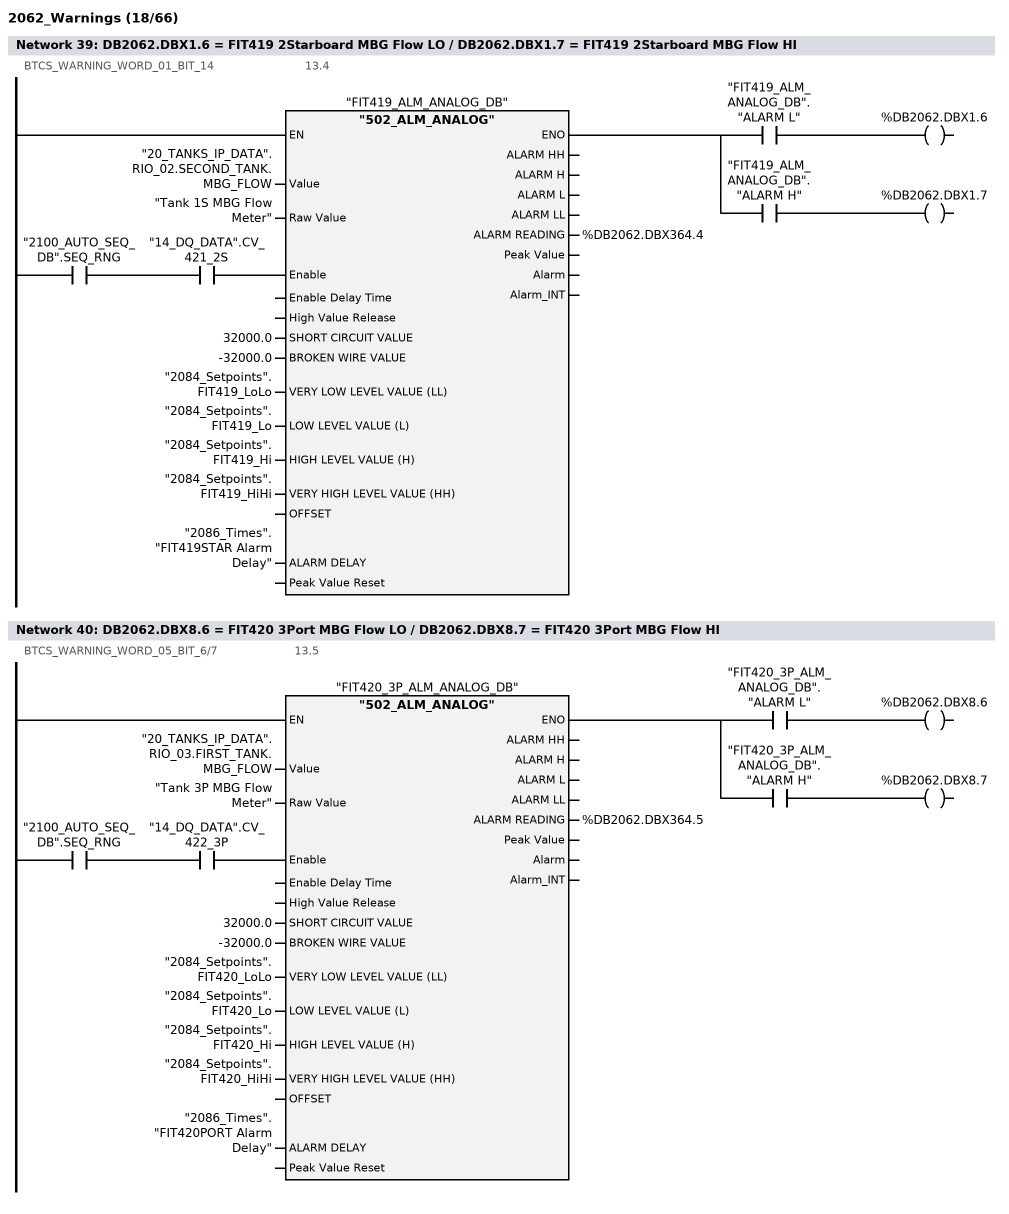
   RUNG wire#powerrail
      "FIT419_ALM_ANALOG_DB"(Enable := wire#w1, Value := "20_TANKS_IP_DATA".RIO_02.SECOND_TANK.MBG_FLOW, "Raw Value" := "Tank 1S MBG Flow Meter", "Enable Delay Time" :=, "High Value Release" :=, "SHORT CIRCUIT VALUE" := 32000.0, "BROKEN WIRE VALUE" := -32000.0, "VERY LOW LEVEL VALUE (LL)" := "2084_Setpoints".FIT419_LoLo, "LOW LEVEL VALUE (L)" := "2084_Setpoints".FIT419_Lo, "HIGH LEVEL VALUE (H)" := "2084_Setpoints".FIT419_Hi, "VERY HIGH LEVEL VALUE (HH)" := "2084_Setpoints".FIT419_HiHi, OFFSET :=, "ALARM DELAY" := "2086_Times"."FIT419STAR Alarm Delay", "Peak Value Reset" :=, "ALARM HH" =>, "ALARM H" =>, "ALARM L" =>, "ALARM LL" =>, "ALARM READING" => %DB2062.DBX364.4, "Peak Value" =>, Alarm =>, Alarm_INT =>)
      wire#w2
      Contact( "FIT419_ALM_ANALOG_DB"."ALARM L" )
      Coil( %DB2062.DBX1.6 )
   END_RUNG
   RUNG wire#powerrail
      Contact( "2100_AUTO_SEQ_DB".SEQ_RNG )
      Contact( "14_DQ_DATA".CV_421_2S )
   END_RUNG wire#w1
   RUNG wire#w2
      Contact( "FIT419_ALM_ANALOG_DB"."ALARM H" )
      Coil( %DB2062.DBX1.7 )
   END_RUNG
   // the same network as SCL:
   "FIT419_ALM_ANALOG_DB"(Value := "20_TANKS_IP_DATA".RIO_02.SECOND_TANK.MBG_FLOW,   // "502_ALM_ANALOG"
                          "Raw Value" := "Tank 1S MBG Flow Meter",
                          Enable := "2100_AUTO_SEQ_DB".SEQ_RNG AND "14_DQ_DATA".CV_421_2S,
                          "SHORT CIRCUIT VALUE" := 32000.0,
                          "BROKEN WIRE VALUE" := -32000.0,
                          "VERY LOW LEVEL VALUE (LL)" := "2084_Setpoints".FIT419_LoLo,
                          "LOW LEVEL VALUE (L)" := "2084_Setpoints".FIT419_Lo,
                          "HIGH LEVEL VALUE (H)" := "2084_Setpoints".FIT419_Hi,
                          "VERY HIGH LEVEL VALUE (HH)" := "2084_Setpoints".FIT419_HiHi,
                          "ALARM DELAY" := "2086_Times"."FIT419STAR Alarm Delay",
                          "ALARM READING" => %DB2062.DBX364.4,
                          ENO => #_w1);
   %DB2062.DBX1.6 := #_w1 AND "FIT419_ALM_ANALOG_DB"."ALARM L";
   %DB2062.DBX1.7 := #_w1 AND "FIT419_ALM_ANALOG_DB"."ALARM H";
END_REGION

REGION Network 40: DB2062.DBX8.6 = FIT420 3Port MBG Flow LO / DB2062.DBX8.7 = FIT420 3Port MBG Flow HI
   // BTCS_WARNING_WORD_05_BIT_6/7                      13.5
   RUNG wire#powerrail
      "FIT420_3P_ALM_ANALOG_DB"(Enable := wire#w1, Value := "20_TANKS_IP_DATA".RIO_03.FIRST_TANK.MBG_FLOW, "Raw Value" := "Tank 3P MBG Flow Meter", "Enable Delay Time" :=, "High Value Release" :=, "SHORT CIRCUIT VALUE" := 32000.0, "BROKEN WIRE VALUE" := -32000.0, "VERY LOW LEVEL VALUE (LL)" := "2084_Setpoints".FIT420_LoLo, "LOW LEVEL VALUE (L)" := "2084_Setpoints".FIT420_Lo, "HIGH LEVEL VALUE (H)" := "2084_Setpoints".FIT420_Hi, "VERY HIGH LEVEL VALUE (HH)" := "2084_Setpoints".FIT420_HiHi, OFFSET :=, "ALARM DELAY" := "2086_Times"."FIT420PORT Alarm Delay", "Peak Value Reset" :=, "ALARM HH" =>, "ALARM H" =>, "ALARM L" =>, "ALARM LL" =>, "ALARM READING" => %DB2062.DBX364.5, "Peak Value" =>, Alarm =>, Alarm_INT =>)
      wire#w2
      Contact( "FIT420_3P_ALM_ANALOG_DB"."ALARM L" )
      Coil( %DB2062.DBX8.6 )
   END_RUNG
   RUNG wire#powerrail
      Contact( "2100_AUTO_SEQ_DB".SEQ_RNG )
      Contact( "14_DQ_DATA".CV_422_3P )
   END_RUNG wire#w1
   RUNG wire#w2
      Contact( "FIT420_3P_ALM_ANALOG_DB"."ALARM H" )
      Coil( %DB2062.DBX8.7 )
   END_RUNG
   // the same network as SCL:
   "FIT420_3P_ALM_ANALOG_DB"(Value := "20_TANKS_IP_DATA".RIO_03.FIRST_TANK.MBG_FLOW,   // "502_ALM_ANALOG"
                           "Raw Value" := "Tank 3P MBG Flow Meter",
                           Enable := "2100_AUTO_SEQ_DB".SEQ_RNG AND "14_DQ_DATA".CV_422_3P,
                           "SHORT CIRCUIT VALUE" := 32000.0,
                           "BROKEN WIRE VALUE" := -32000.0,
                           "VERY LOW LEVEL VALUE (LL)" := "2084_Setpoints".FIT420_LoLo,
                           "LOW LEVEL VALUE (L)" := "2084_Setpoints".FIT420_Lo,
                           "HIGH LEVEL VALUE (H)" := "2084_Setpoints".FIT420_Hi,
                           "VERY HIGH LEVEL VALUE (HH)" := "2084_Setpoints".FIT420_HiHi,
                           "ALARM DELAY" := "2086_Times"."FIT420PORT Alarm Delay",
                           "ALARM READING" => %DB2062.DBX364.5,
                           ENO => #_w1);
   %DB2062.DBX8.6 := #_w1 AND "FIT420_3P_ALM_ANALOG_DB"."ALARM L";
   %DB2062.DBX8.7 := #_w1 AND "FIT420_3P_ALM_ANALOG_DB"."ALARM H";
END_REGION

REGION Network 41: DB2062.DBX9.0 = FIT419 3Starboard MBG Flow LO / DB2062.DBX9.1 = FIT419 3Starboard MBG Flow HI
   // BTCS_WARNING_WORD_05_BIT_8/9                13.6
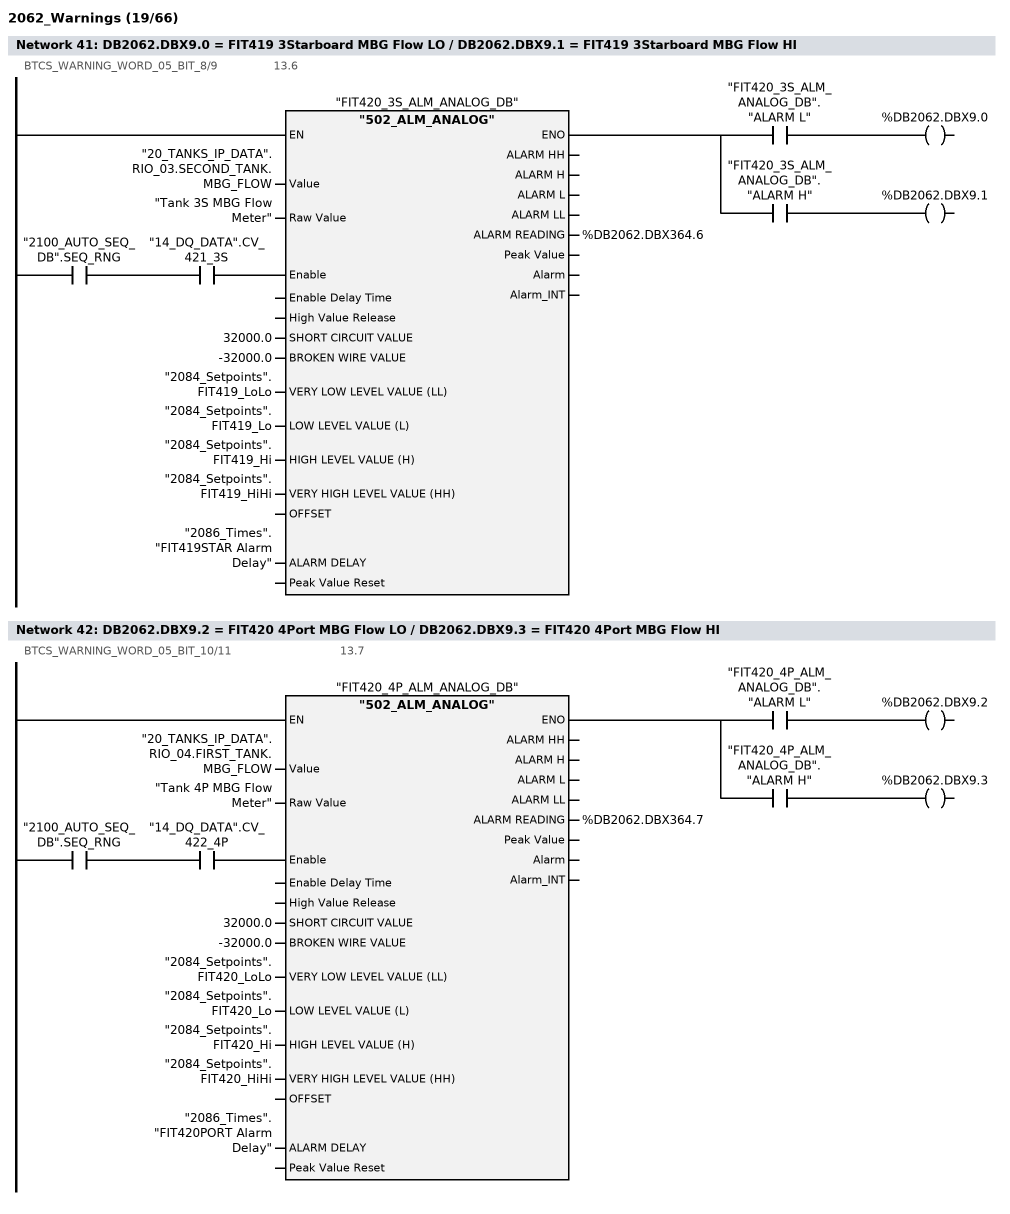
   RUNG wire#powerrail
      "FIT420_3S_ALM_ANALOG_DB"(Enable := wire#w1, Value := "20_TANKS_IP_DATA".RIO_03.SECOND_TANK.MBG_FLOW, "Raw Value" := "Tank 3S MBG Flow Meter", "Enable Delay Time" :=, "High Value Release" :=, "SHORT CIRCUIT VALUE" := 32000.0, "BROKEN WIRE VALUE" := -32000.0, "VERY LOW LEVEL VALUE (LL)" := "2084_Setpoints".FIT419_LoLo, "LOW LEVEL VALUE (L)" := "2084_Setpoints".FIT419_Lo, "HIGH LEVEL VALUE (H)" := "2084_Setpoints".FIT419_Hi, "VERY HIGH LEVEL VALUE (HH)" := "2084_Setpoints".FIT419_HiHi, OFFSET :=, "ALARM DELAY" := "2086_Times"."FIT419STAR Alarm Delay", "Peak Value Reset" :=, "ALARM HH" =>, "ALARM H" =>, "ALARM L" =>, "ALARM LL" =>, "ALARM READING" => %DB2062.DBX364.6, "Peak Value" =>, Alarm =>, Alarm_INT =>)
      wire#w2
      Contact( "FIT420_3S_ALM_ANALOG_DB"."ALARM L" )
      Coil( %DB2062.DBX9.0 )
   END_RUNG
   RUNG wire#powerrail
      Contact( "2100_AUTO_SEQ_DB".SEQ_RNG )
      Contact( "14_DQ_DATA".CV_421_3S )
   END_RUNG wire#w1
   RUNG wire#w2
      Contact( "FIT420_3S_ALM_ANALOG_DB"."ALARM H" )
      Coil( %DB2062.DBX9.1 )
   END_RUNG
   // the same network as SCL:
   "FIT420_3S_ALM_ANALOG_DB"(Value := "20_TANKS_IP_DATA".RIO_03.SECOND_TANK.MBG_FLOW,   // "502_ALM_ANALOG"
                           "Raw Value" := "Tank 3S MBG Flow Meter",
                           Enable := "2100_AUTO_SEQ_DB".SEQ_RNG AND "14_DQ_DATA".CV_421_3S,
                           "SHORT CIRCUIT VALUE" := 32000.0,
                           "BROKEN WIRE VALUE" := -32000.0,
                           "VERY LOW LEVEL VALUE (LL)" := "2084_Setpoints".FIT419_LoLo,
                           "LOW LEVEL VALUE (L)" := "2084_Setpoints".FIT419_Lo,
                           "HIGH LEVEL VALUE (H)" := "2084_Setpoints".FIT419_Hi,
                           "VERY HIGH LEVEL VALUE (HH)" := "2084_Setpoints".FIT419_HiHi,
                           "ALARM DELAY" := "2086_Times"."FIT419STAR Alarm Delay",
                           "ALARM READING" => %DB2062.DBX364.6,
                           ENO => #_w1);
   %DB2062.DBX9.0 := #_w1 AND "FIT420_3S_ALM_ANALOG_DB"."ALARM L";
   %DB2062.DBX9.1 := #_w1 AND "FIT420_3S_ALM_ANALOG_DB"."ALARM H";
END_REGION

REGION Network 42: DB2062.DBX9.2 = FIT420 4Port MBG Flow LO / DB2062.DBX9.3 = FIT420 4Port MBG Flow HI
   // BTCS_WARNING_WORD_05_BIT_10/11                               13.7
   RUNG wire#powerrail
      "FIT420_4P_ALM_ANALOG_DB"(Enable := wire#w1, Value := "20_TANKS_IP_DATA".RIO_04.FIRST_TANK.MBG_FLOW, "Raw Value" := "Tank 4P MBG Flow Meter", "Enable Delay Time" :=, "High Value Release" :=, "SHORT CIRCUIT VALUE" := 32000.0, "BROKEN WIRE VALUE" := -32000.0, "VERY LOW LEVEL VALUE (LL)" := "2084_Setpoints".FIT420_LoLo, "LOW LEVEL VALUE (L)" := "2084_Setpoints".FIT420_Lo, "HIGH LEVEL VALUE (H)" := "2084_Setpoints".FIT420_Hi, "VERY HIGH LEVEL VALUE (HH)" := "2084_Setpoints".FIT420_HiHi, OFFSET :=, "ALARM DELAY" := "2086_Times"."FIT420PORT Alarm Delay", "Peak Value Reset" :=, "ALARM HH" =>, "ALARM H" =>, "ALARM L" =>, "ALARM LL" =>, "ALARM READING" => %DB2062.DBX364.7, "Peak Value" =>, Alarm =>, Alarm_INT =>)
      wire#w2
      Contact( "FIT420_4P_ALM_ANALOG_DB"."ALARM L" )
      Coil( %DB2062.DBX9.2 )
   END_RUNG
   RUNG wire#powerrail
      Contact( "2100_AUTO_SEQ_DB".SEQ_RNG )
      Contact( "14_DQ_DATA".CV_422_4P )
   END_RUNG wire#w1
   RUNG wire#w2
      Contact( "FIT420_4P_ALM_ANALOG_DB"."ALARM H" )
      Coil( %DB2062.DBX9.3 )
   END_RUNG
   // the same network as SCL:
   "FIT420_4P_ALM_ANALOG_DB"(Value := "20_TANKS_IP_DATA".RIO_04.FIRST_TANK.MBG_FLOW,   // "502_ALM_ANALOG"
                           "Raw Value" := "Tank 4P MBG Flow Meter",
                           Enable := "2100_AUTO_SEQ_DB".SEQ_RNG AND "14_DQ_DATA".CV_422_4P,
                           "SHORT CIRCUIT VALUE" := 32000.0,
                           "BROKEN WIRE VALUE" := -32000.0,
                           "VERY LOW LEVEL VALUE (LL)" := "2084_Setpoints".FIT420_LoLo,
                           "LOW LEVEL VALUE (L)" := "2084_Setpoints".FIT420_Lo,
                           "HIGH LEVEL VALUE (H)" := "2084_Setpoints".FIT420_Hi,
                           "VERY HIGH LEVEL VALUE (HH)" := "2084_Setpoints".FIT420_HiHi,
                           "ALARM DELAY" := "2086_Times"."FIT420PORT Alarm Delay",
                           "ALARM READING" => %DB2062.DBX364.7,
                           ENO => #_w1);
   %DB2062.DBX9.2 := #_w1 AND "FIT420_4P_ALM_ANALOG_DB"."ALARM L";
   %DB2062.DBX9.3 := #_w1 AND "FIT420_4P_ALM_ANALOG_DB"."ALARM H";
END_REGION

REGION Network 43: DB2062.DBX9.4 = FIT419 4Starboard MBG Flow LO / DB2062.DBX9.5 = FIT419 4Starboard MBG Flow HI
   // BTCS_WARNING_WORD_05_BIT_12/13                               13.8
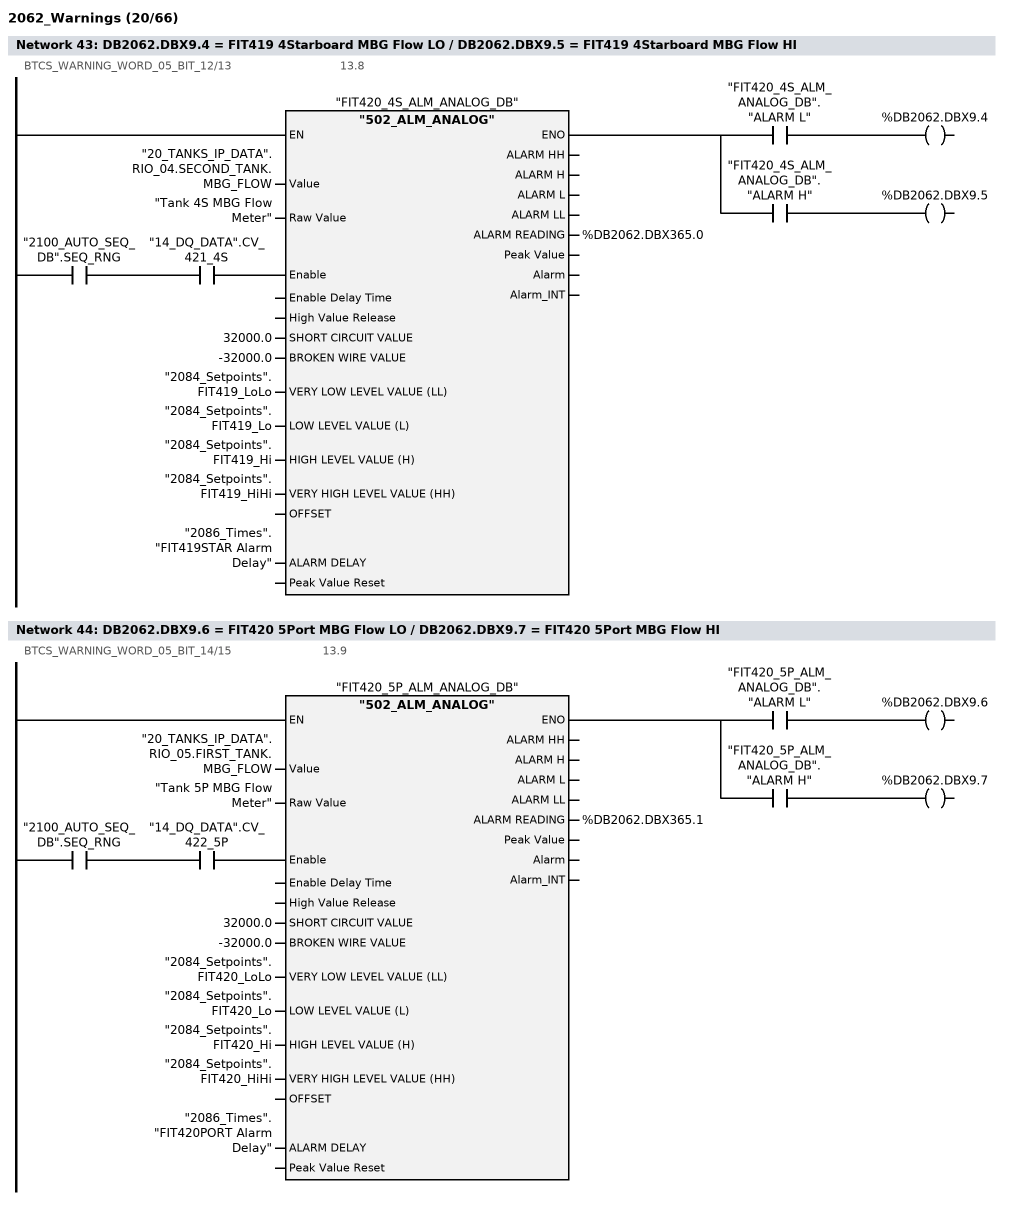
   RUNG wire#powerrail
      "FIT420_4S_ALM_ANALOG_DB"(Enable := wire#w1, Value := "20_TANKS_IP_DATA".RIO_04.SECOND_TANK.MBG_FLOW, "Raw Value" := "Tank 4S MBG Flow Meter", "Enable Delay Time" :=, "High Value Release" :=, "SHORT CIRCUIT VALUE" := 32000.0, "BROKEN WIRE VALUE" := -32000.0, "VERY LOW LEVEL VALUE (LL)" := "2084_Setpoints".FIT419_LoLo, "LOW LEVEL VALUE (L)" := "2084_Setpoints".FIT419_Lo, "HIGH LEVEL VALUE (H)" := "2084_Setpoints".FIT419_Hi, "VERY HIGH LEVEL VALUE (HH)" := "2084_Setpoints".FIT419_HiHi, OFFSET :=, "ALARM DELAY" := "2086_Times"."FIT419STAR Alarm Delay", "Peak Value Reset" :=, "ALARM HH" =>, "ALARM H" =>, "ALARM L" =>, "ALARM LL" =>, "ALARM READING" => %DB2062.DBX365.0, "Peak Value" =>, Alarm =>, Alarm_INT =>)
      wire#w2
      Contact( "FIT420_4S_ALM_ANALOG_DB"."ALARM L" )
      Coil( %DB2062.DBX9.4 )
   END_RUNG
   RUNG wire#powerrail
      Contact( "2100_AUTO_SEQ_DB".SEQ_RNG )
      Contact( "14_DQ_DATA".CV_421_4S )
   END_RUNG wire#w1
   RUNG wire#w2
      Contact( "FIT420_4S_ALM_ANALOG_DB"."ALARM H" )
      Coil( %DB2062.DBX9.5 )
   END_RUNG
   // the same network as SCL:
   "FIT420_4S_ALM_ANALOG_DB"(Value := "20_TANKS_IP_DATA".RIO_04.SECOND_TANK.MBG_FLOW,   // "502_ALM_ANALOG"
                           "Raw Value" := "Tank 4S MBG Flow Meter",
                           Enable := "2100_AUTO_SEQ_DB".SEQ_RNG AND "14_DQ_DATA".CV_421_4S,
                           "SHORT CIRCUIT VALUE" := 32000.0,
                           "BROKEN WIRE VALUE" := -32000.0,
                           "VERY LOW LEVEL VALUE (LL)" := "2084_Setpoints".FIT419_LoLo,
                           "LOW LEVEL VALUE (L)" := "2084_Setpoints".FIT419_Lo,
                           "HIGH LEVEL VALUE (H)" := "2084_Setpoints".FIT419_Hi,
                           "VERY HIGH LEVEL VALUE (HH)" := "2084_Setpoints".FIT419_HiHi,
                           "ALARM DELAY" := "2086_Times"."FIT419STAR Alarm Delay",
                           "ALARM READING" => %DB2062.DBX365.0,
                           ENO => #_w1);
   %DB2062.DBX9.4 := #_w1 AND "FIT420_4S_ALM_ANALOG_DB"."ALARM L";
   %DB2062.DBX9.5 := #_w1 AND "FIT420_4S_ALM_ANALOG_DB"."ALARM H";
END_REGION

REGION Network 44: DB2062.DBX9.6 = FIT420 5Port MBG Flow LO / DB2062.DBX9.7 = FIT420 5Port MBG Flow HI
   // BTCS_WARNING_WORD_05_BIT_14/15                          13.9
   RUNG wire#powerrail
      "FIT420_5P_ALM_ANALOG_DB"(Enable := wire#w1, Value := "20_TANKS_IP_DATA".RIO_05.FIRST_TANK.MBG_FLOW, "Raw Value" := "Tank 5P MBG Flow Meter", "Enable Delay Time" :=, "High Value Release" :=, "SHORT CIRCUIT VALUE" := 32000.0, "BROKEN WIRE VALUE" := -32000.0, "VERY LOW LEVEL VALUE (LL)" := "2084_Setpoints".FIT420_LoLo, "LOW LEVEL VALUE (L)" := "2084_Setpoints".FIT420_Lo, "HIGH LEVEL VALUE (H)" := "2084_Setpoints".FIT420_Hi, "VERY HIGH LEVEL VALUE (HH)" := "2084_Setpoints".FIT420_HiHi, OFFSET :=, "ALARM DELAY" := "2086_Times"."FIT420PORT Alarm Delay", "Peak Value Reset" :=, "ALARM HH" =>, "ALARM H" =>, "ALARM L" =>, "ALARM LL" =>, "ALARM READING" => %DB2062.DBX365.1, "Peak Value" =>, Alarm =>, Alarm_INT =>)
      wire#w2
      Contact( "FIT420_5P_ALM_ANALOG_DB"."ALARM L" )
      Coil( %DB2062.DBX9.6 )
   END_RUNG
   RUNG wire#powerrail
      Contact( "2100_AUTO_SEQ_DB".SEQ_RNG )
      Contact( "14_DQ_DATA".CV_422_5P )
   END_RUNG wire#w1
   RUNG wire#w2
      Contact( "FIT420_5P_ALM_ANALOG_DB"."ALARM H" )
      Coil( %DB2062.DBX9.7 )
   END_RUNG
   // the same network as SCL:
   "FIT420_5P_ALM_ANALOG_DB"(Value := "20_TANKS_IP_DATA".RIO_05.FIRST_TANK.MBG_FLOW,   // "502_ALM_ANALOG"
                           "Raw Value" := "Tank 5P MBG Flow Meter",
                           Enable := "2100_AUTO_SEQ_DB".SEQ_RNG AND "14_DQ_DATA".CV_422_5P,
                           "SHORT CIRCUIT VALUE" := 32000.0,
                           "BROKEN WIRE VALUE" := -32000.0,
                           "VERY LOW LEVEL VALUE (LL)" := "2084_Setpoints".FIT420_LoLo,
                           "LOW LEVEL VALUE (L)" := "2084_Setpoints".FIT420_Lo,
                           "HIGH LEVEL VALUE (H)" := "2084_Setpoints".FIT420_Hi,
                           "VERY HIGH LEVEL VALUE (HH)" := "2084_Setpoints".FIT420_HiHi,
                           "ALARM DELAY" := "2086_Times"."FIT420PORT Alarm Delay",
                           "ALARM READING" => %DB2062.DBX365.1,
                           ENO => #_w1);
   %DB2062.DBX9.6 := #_w1 AND "FIT420_5P_ALM_ANALOG_DB"."ALARM L";
   %DB2062.DBX9.7 := #_w1 AND "FIT420_5P_ALM_ANALOG_DB"."ALARM H";
END_REGION

REGION Network 45: DB2062.DBX10.0 = FIT419 5Starboard MBG Flow LO / DB2062.DBX10.1 = FIT419 5Starboard MBG Flow HI
   // BTCS_WARNING_WORD_06_BIT_0/1                         13.10
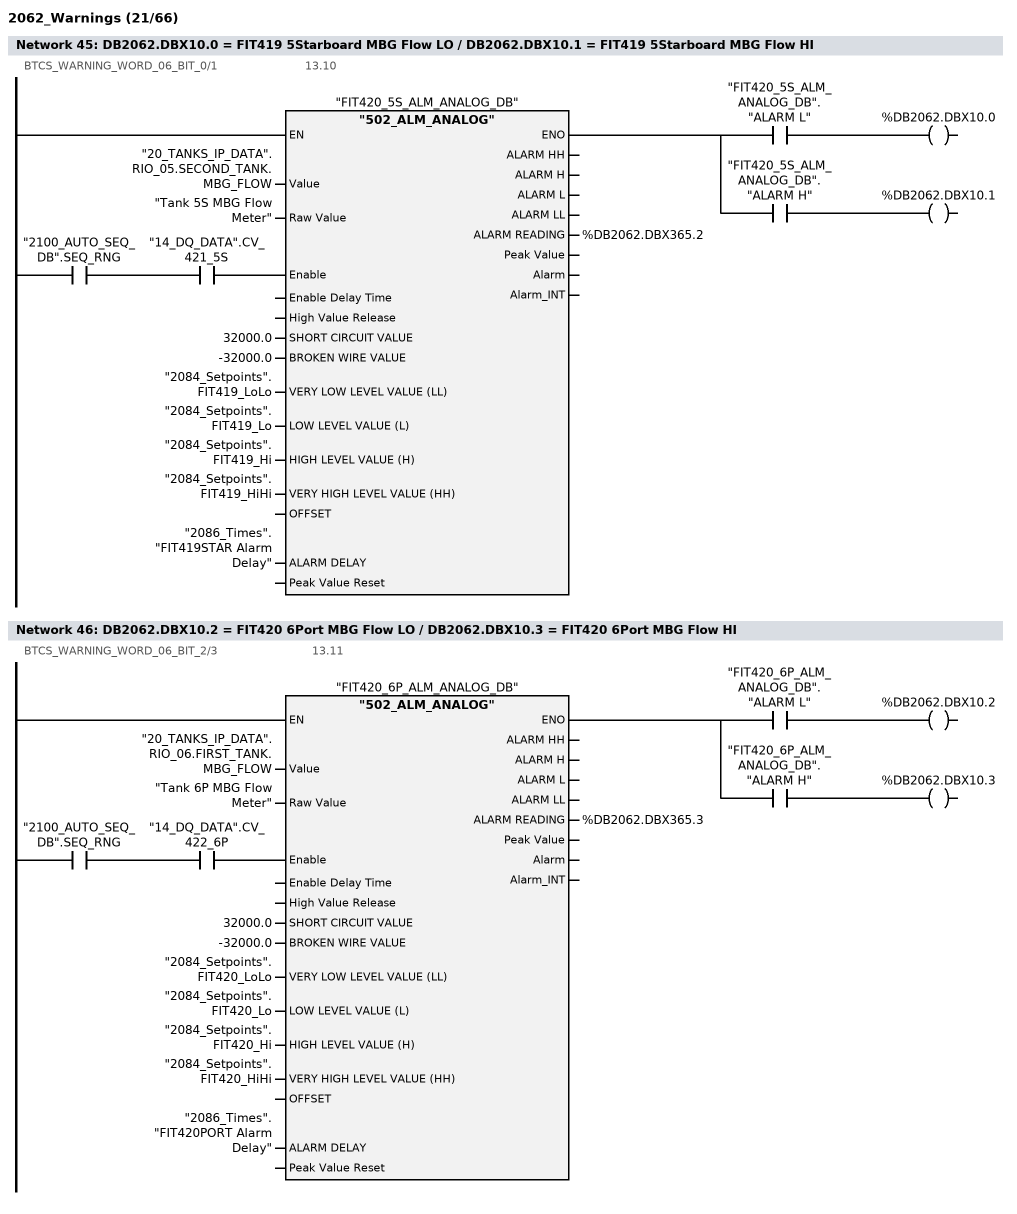
   RUNG wire#powerrail
      "FIT420_5S_ALM_ANALOG_DB"(Enable := wire#w1, Value := "20_TANKS_IP_DATA".RIO_05.SECOND_TANK.MBG_FLOW, "Raw Value" := "Tank 5S MBG Flow Meter", "Enable Delay Time" :=, "High Value Release" :=, "SHORT CIRCUIT VALUE" := 32000.0, "BROKEN WIRE VALUE" := -32000.0, "VERY LOW LEVEL VALUE (LL)" := "2084_Setpoints".FIT419_LoLo, "LOW LEVEL VALUE (L)" := "2084_Setpoints".FIT419_Lo, "HIGH LEVEL VALUE (H)" := "2084_Setpoints".FIT419_Hi, "VERY HIGH LEVEL VALUE (HH)" := "2084_Setpoints".FIT419_HiHi, OFFSET :=, "ALARM DELAY" := "2086_Times"."FIT419STAR Alarm Delay", "Peak Value Reset" :=, "ALARM HH" =>, "ALARM H" =>, "ALARM L" =>, "ALARM LL" =>, "ALARM READING" => %DB2062.DBX365.2, "Peak Value" =>, Alarm =>, Alarm_INT =>)
      wire#w2
      Contact( "FIT420_5S_ALM_ANALOG_DB"."ALARM L" )
      Coil( %DB2062.DBX10.0 )
   END_RUNG
   RUNG wire#powerrail
      Contact( "2100_AUTO_SEQ_DB".SEQ_RNG )
      Contact( "14_DQ_DATA".CV_421_5S )
   END_RUNG wire#w1
   RUNG wire#w2
      Contact( "FIT420_5S_ALM_ANALOG_DB"."ALARM H" )
      Coil( %DB2062.DBX10.1 )
   END_RUNG
   // the same network as SCL:
   "FIT420_5S_ALM_ANALOG_DB"(Value := "20_TANKS_IP_DATA".RIO_05.SECOND_TANK.MBG_FLOW,   // "502_ALM_ANALOG"
                           "Raw Value" := "Tank 5S MBG Flow Meter",
                           Enable := "2100_AUTO_SEQ_DB".SEQ_RNG AND "14_DQ_DATA".CV_421_5S,
                           "SHORT CIRCUIT VALUE" := 32000.0,
                           "BROKEN WIRE VALUE" := -32000.0,
                           "VERY LOW LEVEL VALUE (LL)" := "2084_Setpoints".FIT419_LoLo,
                           "LOW LEVEL VALUE (L)" := "2084_Setpoints".FIT419_Lo,
                           "HIGH LEVEL VALUE (H)" := "2084_Setpoints".FIT419_Hi,
                           "VERY HIGH LEVEL VALUE (HH)" := "2084_Setpoints".FIT419_HiHi,
                           "ALARM DELAY" := "2086_Times"."FIT419STAR Alarm Delay",
                           "ALARM READING" => %DB2062.DBX365.2,
                           ENO => #_w1);
   %DB2062.DBX10.0 := #_w1 AND "FIT420_5S_ALM_ANALOG_DB"."ALARM L";
   %DB2062.DBX10.1 := #_w1 AND "FIT420_5S_ALM_ANALOG_DB"."ALARM H";
END_REGION

REGION Network 46: DB2062.DBX10.2 = FIT420 6Port MBG Flow LO / DB2062.DBX10.3 = FIT420 6Port MBG Flow HI
   // BTCS_WARNING_WORD_06_BIT_2/3                           13.11
   RUNG wire#powerrail
      "FIT420_6P_ALM_ANALOG_DB"(Enable := wire#w1, Value := "20_TANKS_IP_DATA".RIO_06.FIRST_TANK.MBG_FLOW, "Raw Value" := "Tank 6P MBG Flow Meter", "Enable Delay Time" :=, "High Value Release" :=, "SHORT CIRCUIT VALUE" := 32000.0, "BROKEN WIRE VALUE" := -32000.0, "VERY LOW LEVEL VALUE (LL)" := "2084_Setpoints".FIT420_LoLo, "LOW LEVEL VALUE (L)" := "2084_Setpoints".FIT420_Lo, "HIGH LEVEL VALUE (H)" := "2084_Setpoints".FIT420_Hi, "VERY HIGH LEVEL VALUE (HH)" := "2084_Setpoints".FIT420_HiHi, OFFSET :=, "ALARM DELAY" := "2086_Times"."FIT420PORT Alarm Delay", "Peak Value Reset" :=, "ALARM HH" =>, "ALARM H" =>, "ALARM L" =>, "ALARM LL" =>, "ALARM READING" => %DB2062.DBX365.3, "Peak Value" =>, Alarm =>, Alarm_INT =>)
      wire#w2
      Contact( "FIT420_6P_ALM_ANALOG_DB"."ALARM L" )
      Coil( %DB2062.DBX10.2 )
   END_RUNG
   RUNG wire#powerrail
      Contact( "2100_AUTO_SEQ_DB".SEQ_RNG )
      Contact( "14_DQ_DATA".CV_422_6P )
   END_RUNG wire#w1
   RUNG wire#w2
      Contact( "FIT420_6P_ALM_ANALOG_DB"."ALARM H" )
      Coil( %DB2062.DBX10.3 )
   END_RUNG
   // the same network as SCL:
   "FIT420_6P_ALM_ANALOG_DB"(Value := "20_TANKS_IP_DATA".RIO_06.FIRST_TANK.MBG_FLOW,   // "502_ALM_ANALOG"
                           "Raw Value" := "Tank 6P MBG Flow Meter",
                           Enable := "2100_AUTO_SEQ_DB".SEQ_RNG AND "14_DQ_DATA".CV_422_6P,
                           "SHORT CIRCUIT VALUE" := 32000.0,
                           "BROKEN WIRE VALUE" := -32000.0,
                           "VERY LOW LEVEL VALUE (LL)" := "2084_Setpoints".FIT420_LoLo,
                           "LOW LEVEL VALUE (L)" := "2084_Setpoints".FIT420_Lo,
                           "HIGH LEVEL VALUE (H)" := "2084_Setpoints".FIT420_Hi,
                           "VERY HIGH LEVEL VALUE (HH)" := "2084_Setpoints".FIT420_HiHi,
                           "ALARM DELAY" := "2086_Times"."FIT420PORT Alarm Delay",
                           "ALARM READING" => %DB2062.DBX365.3,
                           ENO => #_w1);
   %DB2062.DBX10.2 := #_w1 AND "FIT420_6P_ALM_ANALOG_DB"."ALARM L";
   %DB2062.DBX10.3 := #_w1 AND "FIT420_6P_ALM_ANALOG_DB"."ALARM H";
END_REGION

REGION Network 47: DB2062.DBX10.4 = FIT419 6Starboard MBG Flow LO / DB2062.DBX10.5 = FIT419 6Starboard MBG Flow HI
   // BTCS_WARNING_WORD_06_BIT_4/5                                  13.12
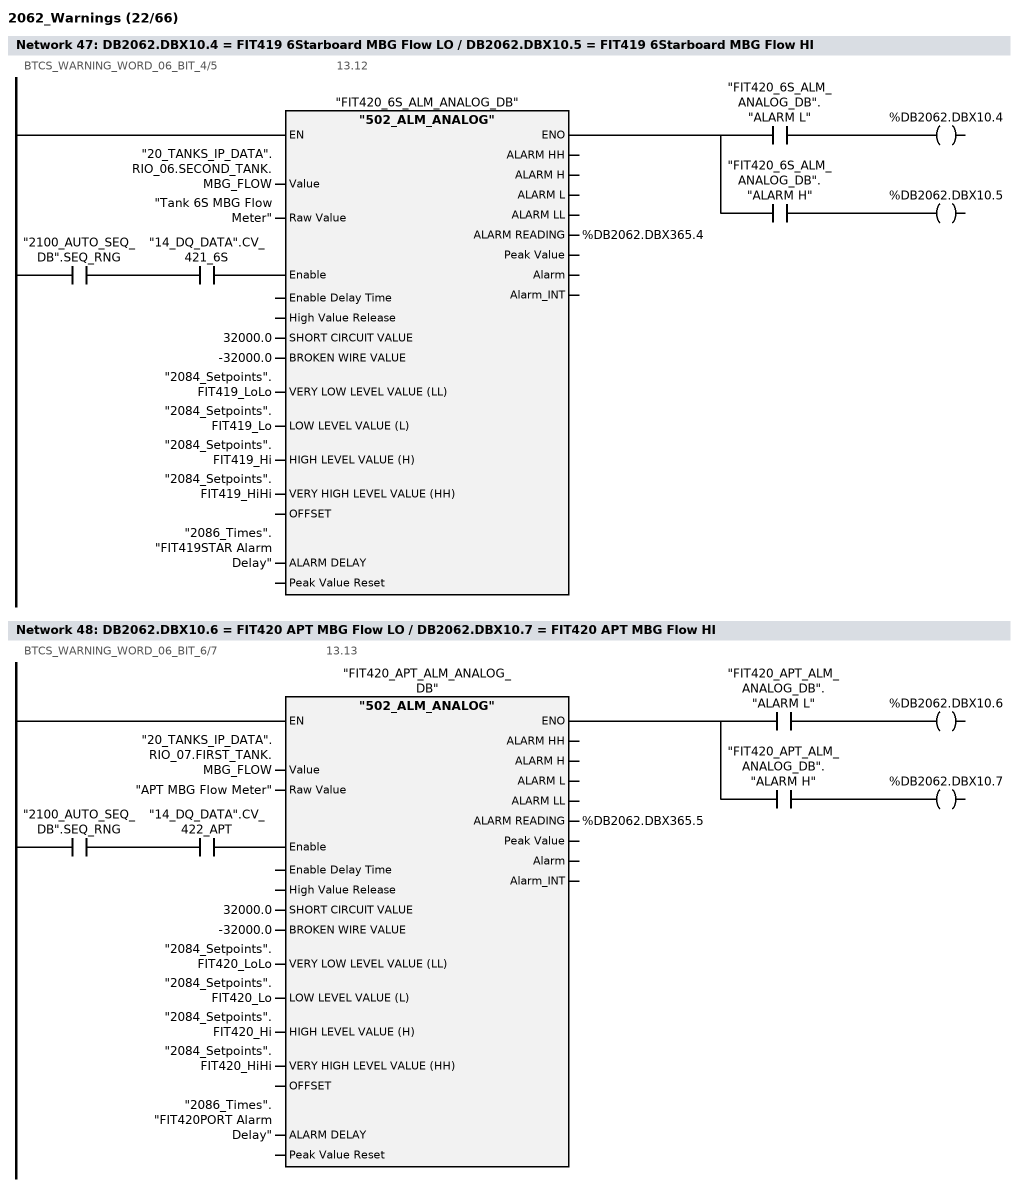
   RUNG wire#powerrail
      "FIT420_6S_ALM_ANALOG_DB"(Enable := wire#w1, Value := "20_TANKS_IP_DATA".RIO_06.SECOND_TANK.MBG_FLOW, "Raw Value" := "Tank 6S MBG Flow Meter", "Enable Delay Time" :=, "High Value Release" :=, "SHORT CIRCUIT VALUE" := 32000.0, "BROKEN WIRE VALUE" := -32000.0, "VERY LOW LEVEL VALUE (LL)" := "2084_Setpoints".FIT419_LoLo, "LOW LEVEL VALUE (L)" := "2084_Setpoints".FIT419_Lo, "HIGH LEVEL VALUE (H)" := "2084_Setpoints".FIT419_Hi, "VERY HIGH LEVEL VALUE (HH)" := "2084_Setpoints".FIT419_HiHi, OFFSET :=, "ALARM DELAY" := "2086_Times"."FIT419STAR Alarm Delay", "Peak Value Reset" :=, "ALARM HH" =>, "ALARM H" =>, "ALARM L" =>, "ALARM LL" =>, "ALARM READING" => %DB2062.DBX365.4, "Peak Value" =>, Alarm =>, Alarm_INT =>)
      wire#w2
      Contact( "FIT420_6S_ALM_ANALOG_DB"."ALARM L" )
      Coil( %DB2062.DBX10.4 )
   END_RUNG
   RUNG wire#powerrail
      Contact( "2100_AUTO_SEQ_DB".SEQ_RNG )
      Contact( "14_DQ_DATA".CV_421_6S )
   END_RUNG wire#w1
   RUNG wire#w2
      Contact( "FIT420_6S_ALM_ANALOG_DB"."ALARM H" )
      Coil( %DB2062.DBX10.5 )
   END_RUNG
   // the same network as SCL:
   "FIT420_6S_ALM_ANALOG_DB"(Value := "20_TANKS_IP_DATA".RIO_06.SECOND_TANK.MBG_FLOW,   // "502_ALM_ANALOG"
                           "Raw Value" := "Tank 6S MBG Flow Meter",
                           Enable := "2100_AUTO_SEQ_DB".SEQ_RNG AND "14_DQ_DATA".CV_421_6S,
                           "SHORT CIRCUIT VALUE" := 32000.0,
                           "BROKEN WIRE VALUE" := -32000.0,
                           "VERY LOW LEVEL VALUE (LL)" := "2084_Setpoints".FIT419_LoLo,
                           "LOW LEVEL VALUE (L)" := "2084_Setpoints".FIT419_Lo,
                           "HIGH LEVEL VALUE (H)" := "2084_Setpoints".FIT419_Hi,
                           "VERY HIGH LEVEL VALUE (HH)" := "2084_Setpoints".FIT419_HiHi,
                           "ALARM DELAY" := "2086_Times"."FIT419STAR Alarm Delay",
                           "ALARM READING" => %DB2062.DBX365.4,
                           ENO => #_w1);
   %DB2062.DBX10.4 := #_w1 AND "FIT420_6S_ALM_ANALOG_DB"."ALARM L";
   %DB2062.DBX10.5 := #_w1 AND "FIT420_6S_ALM_ANALOG_DB"."ALARM H";
END_REGION

REGION Network 48: DB2062.DBX10.6 = FIT420 APT MBG Flow LO / DB2062.DBX10.7 = FIT420 APT MBG Flow HI
   // BTCS_WARNING_WORD_06_BIT_6/7                               13.13
   RUNG wire#powerrail
      "FIT420_APT_ALM_ANALOG_DB"(Enable := wire#w1, Value := "20_TANKS_IP_DATA".RIO_07.FIRST_TANK.MBG_FLOW, "Raw Value" := "APT MBG Flow Meter", "Enable Delay Time" :=, "High Value Release" :=, "SHORT CIRCUIT VALUE" := 32000.0, "BROKEN WIRE VALUE" := -32000.0, "VERY LOW LEVEL VALUE (LL)" := "2084_Setpoints".FIT420_LoLo, "LOW LEVEL VALUE (L)" := "2084_Setpoints".FIT420_Lo, "HIGH LEVEL VALUE (H)" := "2084_Setpoints".FIT420_Hi, "VERY HIGH LEVEL VALUE (HH)" := "2084_Setpoints".FIT420_HiHi, OFFSET :=, "ALARM DELAY" := "2086_Times"."FIT420PORT Alarm Delay", "Peak Value Reset" :=, "ALARM HH" =>, "ALARM H" =>, "ALARM L" =>, "ALARM LL" =>, "ALARM READING" => %DB2062.DBX365.5, "Peak Value" =>, Alarm =>, Alarm_INT =>)
      wire#w2
      Contact( "FIT420_APT_ALM_ANALOG_DB"."ALARM L" )
      Coil( %DB2062.DBX10.6 )
   END_RUNG
   RUNG wire#powerrail
      Contact( "2100_AUTO_SEQ_DB".SEQ_RNG )
      Contact( "14_DQ_DATA".CV_422_APT )
   END_RUNG wire#w1
   RUNG wire#w2
      Contact( "FIT420_APT_ALM_ANALOG_DB"."ALARM H" )
      Coil( %DB2062.DBX10.7 )
   END_RUNG
   // the same network as SCL:
   "FIT420_APT_ALM_ANALOG_DB"(Value := "20_TANKS_IP_DATA".RIO_07.FIRST_TANK.MBG_FLOW,   // "502_ALM_ANALOG"
                           "Raw Value" := "APT MBG Flow Meter",
                           Enable := "2100_AUTO_SEQ_DB".SEQ_RNG AND "14_DQ_DATA".CV_422_APT,
                           "SHORT CIRCUIT VALUE" := 32000.0,
                           "BROKEN WIRE VALUE" := -32000.0,
                           "VERY LOW LEVEL VALUE (LL)" := "2084_Setpoints".FIT420_LoLo,
                           "LOW LEVEL VALUE (L)" := "2084_Setpoints".FIT420_Lo,
                           "HIGH LEVEL VALUE (H)" := "2084_Setpoints".FIT420_Hi,
                           "VERY HIGH LEVEL VALUE (HH)" := "2084_Setpoints".FIT420_HiHi,
                           "ALARM DELAY" := "2086_Times"."FIT420PORT Alarm Delay",
                           "ALARM READING" => %DB2062.DBX365.5,
                           ENO => #_w1);
   %DB2062.DBX10.6 := #_w1 AND "FIT420_APT_ALM_ANALOG_DB"."ALARM L";
   %DB2062.DBX10.7 := #_w1 AND "FIT420_APT_ALM_ANALOG_DB"."ALARM H";
END_REGION

REGION Network 50: DB2062.DBX11.0 = PT415 RIO1 Deck IG Pressure LO / DB2062.DBX11.1 = PT415 RIO1 Deck IG Pressure HI
   // BTCS_WARNING_WORD_06_BIT_8/9                                13.14
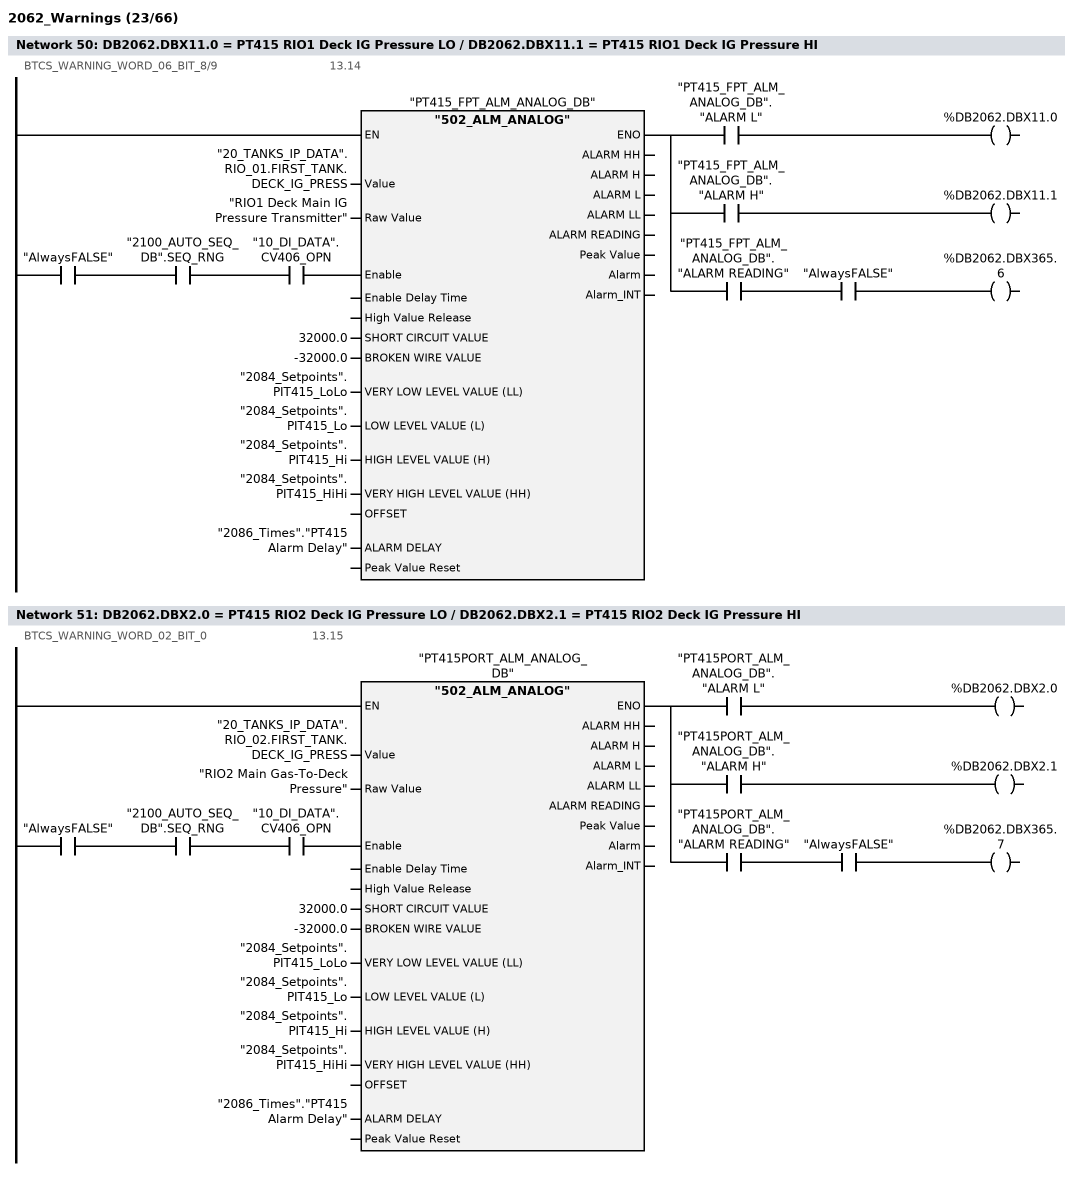
   RUNG wire#powerrail
      "PT415_FPT_ALM_ANALOG_DB"(Enable := wire#w1, Value := "20_TANKS_IP_DATA".RIO_01.FIRST_TANK.DECK_IG_PRESS, "Raw Value" := "RIO1 Deck Main IG Pressure Transmitter", "Enable Delay Time" :=, "High Value Release" :=, "SHORT CIRCUIT VALUE" := 32000.0, "BROKEN WIRE VALUE" := -32000.0, "VERY LOW LEVEL VALUE (LL)" := "2084_Setpoints".PIT415_LoLo, "LOW LEVEL VALUE (L)" := "2084_Setpoints".PIT415_Lo, "HIGH LEVEL VALUE (H)" := "2084_Setpoints".PIT415_Hi, "VERY HIGH LEVEL VALUE (HH)" := "2084_Setpoints".PIT415_HiHi, OFFSET :=, "ALARM DELAY" := "2086_Times"."PT415 Alarm Delay", "Peak Value Reset" :=, "ALARM HH" =>, "ALARM H" =>, "ALARM L" =>, "ALARM LL" =>, "ALARM READING" =>, "Peak Value" =>, Alarm =>, Alarm_INT =>)
      wire#w2
      Contact( "PT415_FPT_ALM_ANALOG_DB"."ALARM L" )
      Coil( %DB2062.DBX11.0 )
   END_RUNG
   RUNG wire#powerrail
      Contact( "AlwaysFALSE" )
      Contact( "2100_AUTO_SEQ_DB".SEQ_RNG )
      Contact( "10_DI_DATA".CV406_OPN )
   END_RUNG wire#w1
   RUNG wire#w2
      Contact( "PT415_FPT_ALM_ANALOG_DB"."ALARM H" )
      Coil( %DB2062.DBX11.1 )
   END_RUNG
   RUNG wire#w2
      Contact( "PT415_FPT_ALM_ANALOG_DB"."ALARM READING" )
      Contact( "AlwaysFALSE" )
      Coil( %DB2062.DBX365.6 )
   END_RUNG
   // the same network as SCL:
   "PT415_FPT_ALM_ANALOG_DB"(Value := "20_TANKS_IP_DATA".RIO_01.FIRST_TANK.DECK_IG_PRESS,   // "502_ALM_ANALOG"
                           "Raw Value" := "RIO1 Deck Main IG Pressure Transmitter",
                           Enable := "AlwaysFALSE" AND "2100_AUTO_SEQ_DB".SEQ_RNG AND "10_DI_DATA".CV406_OPN,
                           "SHORT CIRCUIT VALUE" := 32000.0,
                           "BROKEN WIRE VALUE" := -32000.0,
                           "VERY LOW LEVEL VALUE (LL)" := "2084_Setpoints".PIT415_LoLo,
                           "LOW LEVEL VALUE (L)" := "2084_Setpoints".PIT415_Lo,
                           "HIGH LEVEL VALUE (H)" := "2084_Setpoints".PIT415_Hi,
                           "VERY HIGH LEVEL VALUE (HH)" := "2084_Setpoints".PIT415_HiHi,
                           "ALARM DELAY" := "2086_Times"."PT415 Alarm Delay",
                           ENO => #_w1);
   %DB2062.DBX11.0 := #_w1 AND "PT415_FPT_ALM_ANALOG_DB"."ALARM L";
   %DB2062.DBX11.1 := #_w1 AND "PT415_FPT_ALM_ANALOG_DB"."ALARM H";
   %DB2062.DBX365.6 := #_w1 AND "PT415_FPT_ALM_ANALOG_DB"."ALARM READING" AND "AlwaysFALSE";
END_REGION

REGION Network 51: DB2062.DBX2.0 = PT415 RIO2 Deck IG Pressure LO / DB2062.DBX2.1 = PT415 RIO2 Deck IG Pressure HI
   // BTCS_WARNING_WORD_02_BIT_0                              13.15
   RUNG wire#powerrail
      "PT415PORT_ALM_ANALOG_DB"(Enable := wire#w1, Value := "20_TANKS_IP_DATA".RIO_02.FIRST_TANK.DECK_IG_PRESS, "Raw Value" := "RIO2 Main Gas-To-Deck Pressure", "Enable Delay Time" :=, "High Value Release" :=, "SHORT CIRCUIT VALUE" := 32000.0, "BROKEN WIRE VALUE" := -32000.0, "VERY LOW LEVEL VALUE (LL)" := "2084_Setpoints".PIT415_LoLo, "LOW LEVEL VALUE (L)" := "2084_Setpoints".PIT415_Lo, "HIGH LEVEL VALUE (H)" := "2084_Setpoints".PIT415_Hi, "VERY HIGH LEVEL VALUE (HH)" := "2084_Setpoints".PIT415_HiHi, OFFSET :=, "ALARM DELAY" := "2086_Times"."PT415 Alarm Delay", "Peak Value Reset" :=, "ALARM HH" =>, "ALARM H" =>, "ALARM L" =>, "ALARM LL" =>, "ALARM READING" =>, "Peak Value" =>, Alarm =>, Alarm_INT =>)
      wire#w2
      Contact( "PT415PORT_ALM_ANALOG_DB"."ALARM L" )
      Coil( %DB2062.DBX2.0 )
   END_RUNG
   RUNG wire#powerrail
      Contact( "AlwaysFALSE" )
      Contact( "2100_AUTO_SEQ_DB".SEQ_RNG )
      Contact( "10_DI_DATA".CV406_OPN )
   END_RUNG wire#w1
   RUNG wire#w2
      Contact( "PT415PORT_ALM_ANALOG_DB"."ALARM H" )
      Coil( %DB2062.DBX2.1 )
   END_RUNG
   RUNG wire#w2
      Contact( "PT415PORT_ALM_ANALOG_DB"."ALARM READING" )
      Contact( "AlwaysFALSE" )
      Coil( %DB2062.DBX365.7 )
   END_RUNG
   // the same network as SCL:
   "PT415PORT_ALM_ANALOG_DB"(Value := "20_TANKS_IP_DATA".RIO_02.FIRST_TANK.DECK_IG_PRESS,   // "502_ALM_ANALOG"
                           "Raw Value" := "RIO2 Main Gas-To-Deck Pressure",
                           Enable := "AlwaysFALSE" AND "2100_AUTO_SEQ_DB".SEQ_RNG AND "10_DI_DATA".CV406_OPN,
                           "SHORT CIRCUIT VALUE" := 32000.0,
                           "BROKEN WIRE VALUE" := -32000.0,
                           "VERY LOW LEVEL VALUE (LL)" := "2084_Setpoints".PIT415_LoLo,
                           "LOW LEVEL VALUE (L)" := "2084_Setpoints".PIT415_Lo,
                           "HIGH LEVEL VALUE (H)" := "2084_Setpoints".PIT415_Hi,
                           "VERY HIGH LEVEL VALUE (HH)" := "2084_Setpoints".PIT415_HiHi,
                           "ALARM DELAY" := "2086_Times"."PT415 Alarm Delay",
                           ENO => #_w1);
   %DB2062.DBX2.0 := #_w1 AND "PT415PORT_ALM_ANALOG_DB"."ALARM L";
   %DB2062.DBX2.1 := #_w1 AND "PT415PORT_ALM_ANALOG_DB"."ALARM H";
   %DB2062.DBX365.7 := #_w1 AND "PT415PORT_ALM_ANALOG_DB"."ALARM READING" AND "AlwaysFALSE";
END_REGION

REGION Network 52: DB2062.DBX11.2 = PT415 RIO3 Deck IG Pressure LO / DB2062.DBX11.3 = PT415 RIO3 Deck IG Pressure HI
   // BTCS_WARNING_WORD_06_BIT_10/11                         14.0